screen "0017_Home Screen" 1280x800, template "Navigation"
   on GenerateScreen: SetTag("NavScreenChange", 7)
   on ClearScreen: SetTag("NavScreenChange", 0)
   GraphicView "Alarm Indicator Pump1" at 416,472 size 25x21; Picture "AlarmState2"
      Visibility <- "DB613_Komponent_State_GroupStatus{1}_FaultExist"
   GraphicView "Alarm Indicator Pump2" at 584,472 size 25x21; Picture "AlarmState2"
      Visibility <- "DB613_Komponent_State_GroupStatus{2}_FaultExist"
   GraphicView "Alarm Indicator hydraulic" at 1105,597 size 25x21; Picture "AlarmState2"
      Visibility <- "DB611_Hydraulic_State_MH_Hydraulic{1}_Fault_Exist"
   GraphicView "Alarm Indicator Pump2_1" at 508,688 size 25x21; Picture "AlarmState2"
      Visibility <- "DB614_MH_State_FaulExist"
   Button "Button_25" at 377,130 size 153x214; TextOff 'Text'; PictureOff "motor2"
      on Press: ActivateScreen("0006_Tank", 0); SetTag("DB612_Tank_State.ReadDeviceNo", 1); SetTag("NavScreenChange", 0)
   Button "Button_26" at 537,130 size 153x214; TextOff 'Text'; PictureOff "motor2"
      on Press: ActivateScreen("0006_Tank", 0); SetTag("DB612_Tank_State.ReadDeviceNo", 2); SetTag("NavScreenChange", 0)
   Button "b_Pump1" at 407,466 size 56x48; TextOff 'Text'
      on Press: ActivateScreen("0024_ActualFaults", 0); SetTag("Alarm_Filter_Tag", 3)
      ObjectEnable <- "DB613_Komponent_State_GroupStatus{1}_FaultExist"
   Button "b_Pump2" at 574,466 size 56x48; TextOff 'Text'
      ObjectEnable <- "DB613_Komponent_State_GroupStatus{2}_FaultExist"
      on Press: ActivateScreen("0024_ActualFaults", 0); SetTag("Alarm_Filter_Tag", 3); SetTag("NavScreenChange", 0)
   Button "b_hydraulic" at 1096,592 size 56x48; TextOff 'Text'
      on Press: ActivateScreen("0024_ActualFaults", 0); SetTag("Alarm_Filter_Tag", 2); SetTag("NavScreenChange", 0)
      ObjectEnable <- "DB611_Hydraulic_State_MH_Hydraulic{1}_Fault_Exist"
   Button "b_Pump2_1" at 494,677 size 56x48; TextOff 'Text'
      on Press: ActivateScreen("0024_ActualFaults", 0); SetTag("Alarm_Filter_Tag", 1); SetTag("NavScreenChange", 0)
      ObjectEnable <- "DB614_MH_State_FaulExist"
      Visibility <- "DB614_MH_State_FaulExist"
   GraphicView "Alarm Indicator Tank1" at 444,213 size 25x21; Picture "AlarmState2"
      Visibility <- "DB612_Tank_State_FaultExists{1}"
   GraphicView "Alarm Indicator Tank2" at 602,209 size 25x21; Picture "AlarmState2"
      Visibility <- "DB612_Tank_State_FaultExists{2}"
   Button "b_Tank1" at 432,208 size 50x36; TextOff 'Text'
      ObjectEnable <- "DB612_Tank_State_FaultExists{1}"
      on Press: ActivateScreen("0024_ActualFaults", 0); SetTag("Alarm_Filter_Tag", 4); SetTag("NavScreenChange", 0)
   Button "b_Tank2" at 588,208 size 50x36; TextOff 'Text'
      on Press: ActivateScreen("0024_ActualFaults", 0); SetTag("Alarm_Filter_Tag", 4); SetTag("NavScreenChange", 0)
      ObjectEnable <- "DB612_Tank_State_FaultExists{2}"
   TextField "Text field_8" at 549,392 size 129x30; Text '%'
      Visibility <- "DB702_Tank_Value_Tank{2}_With_Level_Probe"
   TextField "Text field_3" at 549,357 size 129x30; Text 'ºC'
   TextField "Text field_10" at 548,590 size 129x30; Text '%'
   TextField "Text field_14" at 548,526 size 129x30; Text 'bar'
   TextField "Text field_12" at 548,558 size 129x30; Text 'g/s'
   TextField "Text field_15" at 389,526 size 129x30; Text 'bar'
   TextField "Text field_9" at 389,590 size 129x30; Text '%'
   TextField "Text field_13" at 389,558 size 129x30; Text 'g/s'
   TextField "Text field_16" at 501,754 size 95x33; Text 'NL'
      Visibility <- "DB704_MH_Value_Mixinghead{0}_WithInerting"
   TextField "Text field_7" at 389,392 size 129x30; Text '%'
      Visibility <- "DB702_Tank_Value_Tank{1}_With_Level_Probe"
   TextField "Text field_4" at 389,357 size 129x30; Text 'ºC'
   TextField "Text field_2" at 595,640 size 95x33; Text 'bar'
   TextField "Text field_1" at 594,677 size 95x33; Text 'ºC'
   TextField "Text field_6" at 375,677 size 95x33; Text 'ºC'
   IOField "I/O field_20" at 501,754 size 73x33; FormatPattern 9999.9
      ProcessValue <- "DB619_State_MPart_ActMHInerting{1}_Total_Flow_N2_Visu"
      Visibility <- "DB704_MH_Value_Mixinghead{0}_WithInerting"
   IOField "I/O field_11" at 389,357 size 93x30; FormatPattern 9999.9
      ProcessValue <- "DB602_PV_Tank_Tank{1}_Temp_PV_ActV_Value"
   IOField "I/O field_12" at 549,357 size 93x30; FormatPattern 9999.9
      ProcessValue <- "DB602_PV_Tank_Tank{2}_Temp_PV_ActV_Value"
   IOField "I/O field_3" at 595,640 size 73x33; FormatPattern 9999.9
      ProcessValue <- "DB619_State_MPart_ActMHPressureMa{1}_Comp{2}"
   GraphicView "Graphic view_1" at 387,128 size 129x217; Picture "tank"
   GraphicView "Graphic view_2" at 549,128 size 129x217; Picture "tank"
   Button "Button_19" at 391,468 size 121x46; TextOff 'Text'; PictureOff "motor"
      on Click: SetTag("DB613_Komponent_State_ReadDeviceNo", 1); SetTag("NavScreenChange", 0); ActivateScreen("0010_Pump", 0)
   Button "Button_20" at 552,468 size 121x46; TextOff 'Text'; PictureOff "motor2"
      on Click: SetTag("DB613_Komponent_State_ReadDeviceNo", 2); SetTag("NavScreenChange", 0); ActivateScreen("0010_Pump", 0)
   Button "Button_22" at 987,418 size 162x134; TextOff 'MACHINE'; PictureOff "Machine"
      on Press: ActivateScreen("0021_Machine", 0); SetTag("NavScreenChange", 0)
   IOField "I/O field_43" at 378,97 size 151x30; FormatPattern ????????????????????
      ProcessValue <- "DB702_Tank_Value_Tank{1}_Name"
      Appearance <- "DB702_Tank_Value_Tank{1}_Color"
   IOField "I/O field_13" at 538,97 size 151x30; FormatPattern ????????????????????
      Appearance <- "DB702_Tank_Value_Tank{2}_Color"
      ProcessValue <- "DB702_Tank_Value_Tank{2}_Name"
   IOField "I/O field_14" at 378,426 size 151x30; FormatPattern ????????????????????
      Appearance <- "DB702_Tank_Value_Tank{1}_Color"
      ProcessValue <- "DB753_MeteringPump_Pump{1}_Name"
   IOField "I/O field_15" at 538,426 size 151x30; FormatPattern ????????????????????
      Appearance <- "DB702_Tank_Value_Tank{2}_Color"
      ProcessValue <- "DB753_MeteringPump_Pump{2}_Name"
   IOField "I/O field_16" at 703,651 size 151x30; FormatPattern ????????????????????
      Appearance <- "DB702_Tank_Value_Tank{2}_Color"
      ProcessValue <- "DB753_MeteringPump_Pump{2}_Name"
   IOField "I/O field_17" at 212,651 size 151x30; FormatPattern ????????????????????
      ProcessValue <- "DB753_MeteringPump_Pump{1}_Name"
      Appearance <- "DB702_Tank_Value_Tank{1}_Color"
   Button "Button_3" at 1015,579 size 139x135; TextOff 'MH hydrlc'; PictureOff "Mcn"
      on Press: ActivateScreen("0002_MixingHeadHydraulic", 0); SetTag("NavScreenChange", 0)
   TextField "Text field_11" at 459,754 size 41x33; Text 'N2'
      Visibility <- "DB704_MH_Value_Mixinghead{0}_WithInerting"
   GraphicView "Graphic view_3" at 478,640 size 104x112; Picture "images_4"
   GraphicView "Graphic view_5" at 483,637 size 28x27; Picture "cp2"
      Visibility <- "DB614_MH_State_MH_CleaningPiston{0}_Switch_CP_Forward"
   Bar "Bar_2" at 598,166 size 33x142; MinimumValue 0; MaximumValue 100
      ProcessValue <- "DB602_PV_Tank_Tank{2}_Level_PV_ActV_Value"
   TextField "Text field_5" at 375,640 size 95x33; Text 'bar'
   IOField "I/O field_4" at 376,677 size 73x33; FormatPattern 9999.9
      ProcessValue <- "DB619_State_MPart_ActMHTemperatureMa{1}_Comp{1}"
   IOField "I/O field_18" at 389,392 size 93x30; FormatPattern 9999.9
      ProcessValue <- "DB602_PV_Tank_Tank{1}_Level_PV_ActV_Value"
      Visibility <- "DB702_Tank_Value_Tank{1}_With_Level_Probe"
   IOField "I/O field_1" at 594,677 size 73x33; FormatPattern 9999.9
      ProcessValue <- "DB619_State_MPart_ActMHTemperatureMa{1}_Comp{2}"
   IOField "I/O field_19" at 549,392 size 93x30; FormatPattern 9999.9
      ProcessValue <- "DB602_PV_Tank_Tank{2}_Level_PV_ActV_Value"
      Visibility <- "DB702_Tank_Value_Tank{2}_With_Level_Probe"
   IOField "I/O field_5" at 389,526 size 97x30; FormatPattern 9999.9
      ProcessValue <- "DB608_PV_Metering_Metering{1}_Pressure_PV_ActV_Value"
   IOField "I/O field_7" at 548,526 size 97x30; FormatPattern 9999.9
      ProcessValue <- "DB608_PV_Metering_Metering{2}_Pressure_PV_ActV_Value"
   IOField "I/O field_8" at 548,558 size 97x30; FormatPattern 9999.99
      ProcessValue <- "DB608_PV_Metering_Metering{2}_Flow_PV_ActV_Value"
   IOField "I/O field_6" at 389,558 size 97x30; FormatPattern 9999.99
      ProcessValue <- "DB608_PV_Metering_Metering{1}_Flow_PV_ActV_Value"
   IOField "I/O field_9" at 389,590 size 97x30; FormatPattern 9999.9
      ProcessValue <- "DB608_PV_Metering_Metering{1}_MixingRatio_PV_ActV_Value"
   SymbolicIOField "Symbolic I/O field_1" at 406,718 size 102x33; TextOff '0'; TextOn '1'; TextList "MH_NO"
      ProcessValue <- "DB619_State_MPart_SWU{1}_ActualSWU"
      Visibility <- "DB619_State_MPart_SWU{1}_ActualSWU"
   Button "Button_21" at 479,637 size 104x112; TextOff 'Mixinghead'
      on Click: ActivateScreen("0004_Mixinghead", 0)
   IOField "I/O field_10" at 548,590 size 97x30; FormatPattern 9999.9
      ProcessValue <- "DB608_PV_Metering_Metering{2}_MixingRatio_PV_ActV_Value"
   Button "Button_2" at 543,522 size 140x103; TextOff 'Text'
      on Click: SetTag("DB613_Komponent_State_ReadDeviceNo", 2); SetTag("NavScreenChange", 0); ActivateScreen("0010_Pump", 0)
   Button "Button_1" at 383,522 size 140x102; TextOff 'Text'
      on Click: SetTag("DB613_Komponent_State_ReadDeviceNo", 1); SetTag("NavScreenChange", 0); ActivateScreen("0010_Pump", 0)
   GraphicView "ABB ROBOT" at 965,109 size 198x244; Picture "ABB Robot"
      Visibility <- "DB1901_Config_Robots_Config_Robots{0}_Type_ABB"
   GraphicView "KUKA ROBOT" at 965,109 size 198x244; Picture "Kuka Robot"
      Visibility <- "DB1901_Config_Robots_Config_Robots{0}_Type_Kuka"
   GraphicView "MOTOMAN ROBOT" at 965,109 size 198x244; Picture "Motoman Robot"
      Visibility <- "DB1901_Config_Robots_Config_Robots{0}_Type_Motoman"
   GraphicView "FANUC ROBOT" at 965,109 size 198x244; Picture "Fanuc Robot"
      Visibility <- "DB1901_Config_Robots_Config_Robots{0}_Type_Fanuc"
   Button "Button_27" at 955,97 size 175x267; TextOff 'Robot'
      on Click: ActivateScreen("0034_Robot", 0)
      Visibility <- "DB704_MH_Value_Mixinghead{0}_Conf_IntWithRobot"
   IOField "I/O field_2" at 375,640 size 73x33; FormatPattern 9999.9
      ProcessValue <- "DB619_State_MPart_ActMHPressureMa{1}_Comp{1}"
   Rectangle "Rectangle_8" at 598,166 size 33x142
      Visibility <- "DB612_Tank_State_Tank{2}_Max_Level"
   Rectangle "Rectangle_3" at 598,262 size 33x46
      Visibility <- "DB612_Tank_State_Tank{2}_Min_Level"
   Rectangle "Rectangle_5" at 598,166 size 33x142
      Visibility <- "DB612_Tank_State_Tank{2}_Start_Level_Filling"
   Rectangle "Rectangle_4" at 598,166 size 33x142
      Visibility <- "DB612_Tank_State_Tank{2}_Max_Level"
   Rectangle "Rectangle_7" at 440,166 size 33x142
      Visibility <- "DB612_Tank_State_Tank{1}_Max_Level"
   Rectangle "Rectangle_2" at 440,262 size 33x46
      Visibility <- "DB612_Tank_State_Tank{1}_Min_Level"
   Rectangle "Rectangle_6" at 440,166 size 33x142
      Visibility <- "DB612_Tank_State_Tank{1}_Start_Level_Filling"
   Rectangle "Rectangle_1" at 440,166 size 33x142
      Visibility <- "DB612_Tank_State_Tank{1}_Max_Level"

screen "0002_MixingHeadHydraulic" 1280x800, template "Navigation"
   on GenerateScreen: SetBit("DB611_Hydraulic_State_Read"); SetTag("Navigation_7", 5)
   IOField "I/O field_1" at 782,261 size 81x30; Authorization "Operate"; FormatPattern 99999
      ProcessValue <- "DB721_MH_Hydraulic_MH_Hyd{0}_Hyd_P_Startup"
   IOField "I/O field_2" at 782,293 size 81x30; Authorization "Operate"; FormatPattern 99999
      ProcessValue <- "DB721_MH_Hydraulic_MH_Hyd{0}_Hyd_P_Supervision"
   IOField "I/O field_3" at 782,353 size 81x30; Authorization "Operate"; FormatPattern 99999
      ProcessValue <- "DB721_MH_Hydraulic_MH_Hyd{0}_Hyd_CP_Time"
   IOField "I/O field_4" at 782,385 size 81x30; Authorization "Operate"; FormatPattern 99999
      ProcessValue <- "DB721_MH_Hydraulic_MH_Hyd{0}_Hyd_SwitchOFFDelay"
   IOField "I/O field_5" at 782,417 size 81x30; Authorization "Operate"; FormatPattern 99999
      ProcessValue <- "DB721_MH_Hydraulic_MH_Hyd{0}_Hyd_PressureSwitch"
   IOField "I/O field_6" at 229,521 size 131x30; FormatPattern 9999
      ProcessValue <- "DB611_Hydraulic_State_MH_Hydraulic{0}_HourCounter"
   TextField "Text field_1" at 504,263 size 186x25; Text 'Built up time start:'
   TextField "Text field_2" at 504,295 size 233x25; Text 'Built up time operaring:'
   TextField "Text field_3" at 504,355 size 225x25; Text 'Pressuring time for CP:'
   TextField "Text field_4" at 504,387 size 144x25; Text 'Stand by time:'
   TextField "Text field_5" at 504,419 size 161x25; Text 'Pressuring time:'
   TextField "Text field_6" at 874,263 size 46x25; Text 's'
   TextField "Text field_7" at 874,295 size 46x25; Text 's'
   TextField "Text field_8" at 874,355 size 46x25; Text 's'
   TextField "Text field_9" at 874,387 size 46x25; Text 's'
   TextField "Text field_10" at 874,419 size 46x25; Text 's'
   TextField "Text field_11" at 362,523 size 46x25; Text 'h'
   TextField "Text field_12" at 493,497 size 79x25; Text 'Options'
      Visibility <- "MixingHead Options"
   TextField "Text field_13" at 493,530 size 220x25; Text 'With 2 press switches:'
      Visibility <- "MixingHead Options"
   TextField "Text field_14" at 493,557 size 64x25; Text 'spare:'
      Visibility <- "MixingHead Options"
   TextField "Text field_15" at 493,587 size 64x25; Text 'spare:'
      Visibility <- "MixingHead Options"
   TextField "Text field_16" at 493,617 size 64x25; Text 'spare:'
      Visibility <- "MixingHead Options"
   TextField "Text field_17" at 493,647 size 64x25; Text 'spare:'
      Visibility <- "MixingHead Options"
   GraphicView "Graphic view_4" at 111,179 size 250x272; Picture "Mcn"
   Button "Button_3" at 326,104 size 451x32; TextOff 'MixingHead Hydraulic'
   Button "Button_1" at 482,240 size 423x221; TextOff 'Text'
   Button "Button_2" at 481,468 size 423x220; TextOff 'Text'
      Visibility <- "MixingHead Options"
   Button "check_with_2_press_switch" at 829,527 size 45x30; TextOff 'Text'; PictureOff "download"; PictureList "Check_Uncheck"
      ProcessValue <- "DB721_MH_Hydraulic_Option{0}_With2PSwitch"
      Visibility <- "MixingHead Options"
      on Click: InvertBit("DB721_MH_Hydraulic_Option{0}_With2PSwitch")
   Button "b_Close_MHhydraulic" at 848,470 size 51x41; TextOff 'Text'; PictureOff "images (1)"
      Visibility <- "MixingHead Options"
      on Click: SetTag("MixingHead Options", 0); SetTag("NavScreenChange", 0)
   Button "Button_10" at 1006,248 size 81x116; TextOff 'Text'
   GraphicView "Graphic view_1" at 1019,305 size 55x55; Picture "H"
   Rectangle "Rectangle_1" at 1015,256 size 64x56
      Appearance <- "DB611_Hydraulic_State_MH_Hydraulic{0}_State_Hydraulic"
   GraphicIOField "Graphic I/O field_1" at 1023,260 size 48x48; PictureList "ON_OFF_SWITCH"
      ProcessValue <- "DB611_Hydraulic_State_MH_Hydraulic{0}_Switch_Hydraulic_ON_OFF"
   Button "Button_18" at 1002,240 size 88x128; TextOff 'Text'
      on Click: InvertBit("DB611_Hydraulic_State_MH_Hydraulic{0}_Switch_Hydraulic_ON_OFF")
   GraphicView "Graphic view_2" at 143,508 size 77x51; Picture "counter hydraulic"
   Button "Button_4" at 217,210 size 80x52; TextOff 'Text'
   GraphicView "Graphic view_3" at 250,224 size 25x25; Picture "AlarmState2"
      Visibility <- "DB611_Hydraulic_State_MH_Hydraulic{0}_Fault_Exist"
   Button "b_MH_Increase" at 789,104 size 46x32; TextOff 'Text'; PictureOff "right arrow"
   Button "b_MH_Decrease" at 267,104 size 46x32; TextOff 'Text'; PictureOff "left arrow"
   Button "Template_Button_41" at 16,724 size 68x66; TextOff 'Text'; PictureList "Ico_navigation_2"; PictureOff "Setting_Nav_7"; Authorization "User administration"
      ProcessValue <- "Nav_7"
      Visibility <- "NavUserChange"
      on Click: SetTag("MixingHead Options", 1)

screen "0024_ActualFaults" 1280x800, template "Navigation"
   on ClearScreen: SetTag("refresh_Alarm", 0); SetTag("NavScreenChange", 0)
   on GenerateScreen: SetTag("NavScreenChange", 1)
   AlarmView "Machine Display alarm" at 103,169 size 1072x522
      Visibility <- "Alarm_Filter_Tag"
   Button "Button_3" at 326,104 size 451x32; TextOff 'Actual Fault'; TextList "Alarm_Screen_Filter"
      ProcessValue <- "Alarm_Filter_Tag"
   Button "b_Actual_Alarm" at 1097,92 size 60x60; TextOff 'ACTUAL'; PictureOff "Graphic_28"
      Appearance <- "Alarm_Filter_Tag"
      on Press: SetTag("Alarm_Filter_Tag", 0)
   Button "b_ArchiveAlarm" at 1028,91 size 60x60; TextOff 'ARCHIV'; PictureOff "archiveFoam_1"
      on Click: SetTag("Alarm_Filter_Tag", 10)
      Visibility <- "Alarm_Filter_Tag"
   Button "b_System" at 799,712 size 60x60; TextOff 'System'; PictureOff "system messages"; PictureList "ico_System_message_2"
      Visibility <- "Alarm_Filter_Tag"
      Appearance <- "Alarm_Filter_Tag"
      on Click: SetTag("Alarm_Filter_Tag", 13)
      ProcessValue <- "Alarm_Filter_Tag"
   Button "b_Foaming" at 891,712 size 60x60; TextOff 'Foaming'; PictureList "ico_Foaming_2"
      Visibility <- "Alarm_Filter_Tag"
      Appearance <- "Alarm_Filter_Tag"
      on Click: SetTag("Alarm_Filter_Tag", 12)
      ProcessValue <- "Alarm_Filter_Tag"
   Button "b_FaultFoam" at 984,712 size 60x60; TextOff 'Fault/ Foam'; PictureList "ico_ActualFault_Foaming_2"
      on Click: SetTag("Alarm_Filter_Tag", 10)
      Visibility <- "Alarm_Filter_Tag"
      Appearance <- "Alarm_Filter_Tag"
      ProcessValue <- "Alarm_Filter_Tag"
   Button "b_USB" at 705,712 size 60x60; TextOff 'Export USB'; PictureOff "USB_1"
      on Click: function_e9be9208(1, "Schicht0", '\Storage Card USB\', 0)
   Button "b_Fault_1" at 1077,712 size 60x60; TextOff 'Fault'; PictureList "ico_Actual_Fault_2"
      on Click: SetTag("Alarm_Filter_Tag", 11)
      Visibility <- "Alarm_Filter_Tag"
      ProcessValue <- "Alarm_Filter_Tag"
      Appearance <- "Alarm_Filter_Tag"
   Button "b_Fault_2" at 1077,712 size 60x60; TextOff 'Fault'
      on Click: SetTag("Alarm_Filter_Tag", 11)
      Visibility <- "Alarm_Filter_Tag"
      Appearance <- "Alarm_Filter_Tag"
   Button "b_Foaming_1" at 891,712 size 60x60; TextOff 'Foaming'
      on Click: SetTag("Alarm_Filter_Tag", 12)
      Appearance <- "Alarm_Filter_Tag"
      Visibility <- "Alarm_Filter_Tag"
   Button "b_FaultFoam_1" at 984,712 size 60x60; TextOff 'Fault/ Foam'
      on Click: SetTag("Alarm_Filter_Tag", 10)
      Visibility <- "Alarm_Filter_Tag"
      Appearance <- "Alarm_Filter_Tag"
   Button "b_System_1" at 799,712 size 60x60; TextOff 'System'; PictureOff "system messages"
      on Click: SetTag("Alarm_Filter_Tag", 13)
      Appearance <- "Alarm_Filter_Tag"
      Visibility <- "Alarm_Filter_Tag"
   Button "b_ArchiveAlarm_1" at 1028,91 size 60x60; TextOff 'ARCHIV'; PictureOff "archiveFoam_2"
      on Click: SetTag("Alarm_Filter_Tag", 10)
      Visibility <- "Alarm_Filter_Tag"
   AlarmView "MixingHydraulic Display Alarm" at 103,169 size 1072x522
      Visibility <- "Alarm_Filter_Tag"
   AlarmView "Tank Display Alarm" at 103,169 size 1072x522
      Visibility <- "Alarm_Filter_Tag"
   AlarmView "Pump Display Alarm" at 103,169 size 1072x522
      Visibility <- "Alarm_Filter_Tag"
   AlarmView "Archive faults" at 103,169 size 1072x522; AlarmLog "Schicht0"
      Visibility <- "Alarm_Filter_Tag"
   AlarmView "Archive faults/foaming" at 103,169 size 1072x522; AlarmLog "Schicht0"
      Visibility <- "Alarm_Filter_Tag"
   AlarmView "Archive foaming data" at 103,169 size 1072x522; AlarmLog "Schicht0"
      Visibility <- "Alarm_Filter_Tag"
   AlarmView "Archive system message" at 103,169 size 1072x522; AlarmLog "Schicht0"
      Visibility <- "Alarm_Filter_Tag"
   Button "b_Alarm_MHhydraulic_1" at 122,712 size 60x60; TextOff 'Text'; PictureList "icon_MHalarm"
      Visibility <- "Alarm_Filter_Tag"
      ProcessValue <- "Alarm_Filter_Tag"
      Appearance <- "Alarm_Filter_Tag"
   AlarmView "MixingHead Display Alarm" at 103,169 size 1072x522
      Visibility <- "Alarm_Filter_Tag"
   Button "b_Alarm_MH" at 117,704 size 71x77; TextOff 'MH'
      on Press: SetTag("Alarm_Filter_Tag", 1)
      Visibility <- "Alarm_Filter_Tag"
   AlarmView "Current Display Alarm" at 103,169 size 1072x522
      Visibility <- "Alarm_Filter_Tag"
   Button "b_Alarm_MHhydraulic_2" at 210,712 size 60x60; TextOff 'Text'; PictureList "icon_MHhyraulic"
      Visibility <- "Alarm_Filter_Tag"
      Appearance <- "Alarm_Filter_Tag"
      ProcessValue <- "Alarm_Filter_Tag"
   Button "b_Alarm_MHhydraulic" at 205,704 size 71x77; TextOff 'HYDRLC'
      on Press: SetTag("Alarm_Filter_Tag", 2)
      Visibility <- "Alarm_Filter_Tag"
   Button "b_Alarm_MHhydraulic_3" at 297,712 size 60x60; TextOff 'Text'; PictureList "ico_Pump"
      Visibility <- "Alarm_Filter_Tag"
      Appearance <- "Alarm_Filter_Tag"
      ProcessValue <- "Alarm_Filter_Tag"
   Button "b_MH_DosingPump" at 292,704 size 71x77; TextOff 'DOSING'
      on Press: SetTag("Alarm_Filter_Tag", 3)
      Visibility <- "Alarm_Filter_Tag"
   Button "b_Alarm_MHhydraulic_4" at 471,712 size 60x60; TextOff 'Text'; PictureList "ico_machine"
      Visibility <- "Alarm_Filter_Tag"
      Appearance <- "Alarm_Filter_Tag"
      ProcessValue <- "Alarm_Filter_Tag"
   Button "b_Alarm_Machine" at 466,704 size 71x77; TextOff 'MCHN'
      on Press: SetTag("Alarm_Filter_Tag", 5)
      Visibility <- "Alarm_Filter_Tag"
   Button "b_Alarm_MHhydraulic_5" at 384,712 size 60x60; TextOff 'Text'; PictureList "ico_tank"
      Visibility <- "Alarm_Filter_Tag"
      Appearance <- "Alarm_Filter_Tag"
      ProcessValue <- "Alarm_Filter_Tag"
   Button "b_Alarm_Tank" at 379,704 size 71x77; TextOff 'TANK'
      on Press: SetTag("Alarm_Filter_Tag", 4)
      Visibility <- "Alarm_Filter_Tag"

screen "0015_Oscilloscope" 1280x800, template "Navigation"
   Button "Button_3" at 326,104 size 451x32; TextOff 'Oscilloscope'
   TrendView "Trend view_1" at 105,152 size 1067x565
      ValueAxis1Begin <- "DB025_Oszilloskop_SkalierungGraphLinks_Startwert"
      ValueAxis1End <- "DB025_Oszilloskop_SkalierungGraphLinks_Ebdwert"
      ValueAxis2Begin <- "DB025_Oszilloskop_SkalierungGraphRechts_Startwert"
      ValueAxis2End <- "DB025_Oszilloskop_SkalierungGraphRechts_Ebdwert"
   Button "Button_2" at 115,748 size 52x37; TextOff 'Text'; PictureOff "Graphic_32"
      on Click: function_e0f5d53a("Trend view_1")
   Button "Button_4" at 183,748 size 52x37; TextOff 'Text'; PictureOff "Graphic_31"
      on Click: function_e0f5d53a("Trend view_1")
   Button "Button_5" at 252,748 size 52x37; TextOff 'Text'; PictureOff "Graphic_33"
      on Click: function_b4e726f8("Trend view_1")
   Button "Button_6" at 320,748 size 52x37; TextOff 'Text'; PictureOff "Graphic_34"
      on Click: function_f26ff0ec("Trend view_1")
   Button "Button_7" at 389,748 size 52x37; TextOff 'Text'; PictureOff "Graphic_35"
      on Click: function_c2ce674d("Trend view_1")
   Button "Button_8" at 457,748 size 52x37; TextOff 'Text'; PictureOff "Graphic_36"
      on Click: function_f48c2799("Trend view_1")
   Button "Button_9" at 526,748 size 52x37; TextOff 'Text'; PictureOff "Graphic_37"
      on Click: function_b22ecfcd("Trend view_1")
   Button "Button_10" at 595,748 size 52x37; TextOff 'Text'; PictureOff "gear_setting"
      on Click: ActivateScreen("0016_Osciloscope Setting", 0)
   Button "Button_11" at 979,748 size 52x37; TextOff 'Text'; PictureOff "Graphic_38"
      on Click: function_a3fbdc78("Trend view_1")
   Button "Button_1" at 1047,748 size 52x37; TextOff 'Text'; PictureOff "Graphic_39"
      on Click: function_a16a7cb4("Trend view_1")
   Button "Button_12" at 1115,748 size 52x37; TextOff 'Text'; PictureOff "Graphic_40"
      on Click: function_c7513061("Trend view_1")

screen "0100_LargeScalledValues" 1280x800, template "Navigation"
   Button "Button_2" at 115,466 size 1047x206; TextOff 'Text'
      Appearance <- "DB702_Tank_Value_Tank{2}_Color"
      Visibility <- "LargeScalleValues Control"
   IOField "I/O field_4" at 172,488 size 328x166; FormatPattern 999.9
      ProcessValue <- "DB608_PV_Metering_Metering{2}_Pressure_PV_ActV_Value"
      Visibility <- "LargeScalleValues Control"
   Button "Button_1" at 115,255 size 1047x206; TextOff 'Text'
      Appearance <- "DB702_Tank_Value_Tank{1}_Color"
      Visibility <- "LargeScalleValues Control"
   IOField "I/O field_1" at 172,280 size 328x166; FormatPattern 999.9
      ProcessValue <- "DB608_PV_Metering_Metering{1}_Pressure_PV_ActV_Value"
      Visibility <- "LargeScalleValues Control"
   IOField "I/O field_2" at 836,280 size 328x166; FormatPattern 999.9
      ProcessValue <- "DB608_PV_Metering_Metering{1}_Flow_PV_ActV_Value"
      Visibility <- "LargeScalleValues Control"
   IOField "I/O field_3" at 836,488 size 328x166; FormatPattern 999.9
      ProcessValue <- "DB608_PV_Metering_Metering{2}_Flow_PV_ActV_Value"
      Visibility <- "LargeScalleValues Control"
   TextField "Text field_1" at 252,132 size 192x120; Text 'bar'
      Visibility <- "LargeScalleValues Control"
   TextField "Text field_2" at 872,132 size 192x120; Text 'g/s'
      Visibility <- "LargeScalleValues Control"
   Button "Button_4" at 115,466 size 1047x206; TextOff 'Text'
      Appearance <- "DB702_Tank_Value_Tank{2}_Color"
      Visibility <- "LargeScalleValues Control"
   Button "Button_5" at 115,255 size 1047x206; TextOff 'Text'
      Appearance <- "DB702_Tank_Value_Tank{1}_Color"
      Visibility <- "LargeScalleValues Control"
   IOField "I/O field_5" at 479,280 size 328x166; FormatPattern 999.9
      ProcessValue <- "DB602_PV_Tank_Tank{1}_Level_PV_ActV_Value"
      Visibility <- "LargeScalleValues Control"
   IOField "I/O field_6" at 476,494 size 328x166; FormatPattern 999.9
      ProcessValue <- "DB602_PV_Tank_Tank{2}_Level_PV_ActV_Value"
      Visibility <- "LargeScalleValues Control"
   TextField "Text field_3" at 894,308 size 192x120; Text '%'
      Visibility <- "LargeScalleValues Control"
   TextField "Text field_7" at 894,509 size 192x120; Text '%'
      Visibility <- "LargeScalleValues Control"
   Button "Button_6" at 115,466 size 1047x206; TextOff 'Text'
      Visibility <- "LargeScalleValues Control"
      Appearance <- "DB702_Tank_Value_Tank{2}_Color"
   Button "Button_7" at 115,255 size 1047x206; TextOff 'Text'
      Appearance <- "DB702_Tank_Value_Tank{1}_Color"
      Visibility <- "LargeScalleValues Control"
   TextField "Text field_4" at 252,132 size 192x120; Text 'bar'
      Visibility <- "LargeScalleValues Control"
   TextField "Text field_5" at 872,132 size 192x120; Text 'g/s'
      Visibility <- "LargeScalleValues Control"
   IOField "I/O field_7" at 172,280 size 328x166; FormatPattern 999.9
      ProcessValue <- "DB619_State_MPart_ActMHPressureMa{1}_Comp{1}"
      Visibility <- "LargeScalleValues Control"
   IOField "I/O field_8" at 836,280 size 328x166; FormatPattern 999.9
      ProcessValue <- "DB608_PV_Metering_Metering{1}_Flow_PV_ActV_Value"
      Visibility <- "LargeScalleValues Control"
   IOField "I/O field_9" at 836,488 size 328x166; FormatPattern 999.9
      ProcessValue <- "DB608_PV_Metering_Metering{2}_Flow_PV_ActV_Value"
      Appearance <- "DB702_Tank_Value_Tank{2}_Color"
      Visibility <- "LargeScalleValues Control"
   IOField "I/O field_10" at 172,488 size 328x166; FormatPattern 999.9
      ProcessValue <- "DB619_State_MPart_ActMHPressureMa{1}_Comp{2}"
      Visibility <- "LargeScalleValues Control"
   TextField "Text field_6" at 447,132 size 383x120; Text '---'
      Visibility <- "LargeScalleValues Control"
   Button "Button_8" at 135,711 size 60x60; TextOff 'Text'; PictureList "ico_MH"
      Appearance <- "LargeScalleValues Control"
      ProcessValue <- "LargeScalleValues Control"
   Button "Button_3" at 326,104 size 451x32; TextOff 'Large Scalled Values'
   Button "Button_9" at 296,711 size 60x60; TextOff 'Text'; PictureOff "tank"
      Appearance <- "LargeScalleValues Control"
   Button "Button_10" at 216,711 size 60x60; TextOff 'Text'; PictureOff "Graphic_1"; PictureList "ico_Pump_large"
      Appearance <- "LargeScalleValues Control"
      ProcessValue <- "LargeScalleValues Control"
   Button "b_MH_large" at 135,711 size 60x60; TextOff 'MH'; PictureList "MixingHead"
      Appearance <- "LargeScalleValues Control"
      on Click: SetTag("LargeScalleValues Control", 0)
   Button "b_pump_" at 216,711 size 60x60; TextOff 'Tank'; PictureList "tank"
      on Click: SetTag("LargeScalleValues Control", 1)
   Button "b_tank_large_1" at 296,711 size 60x60; TextOff 'Tank'; PictureList "tank"
      on Click: SetTag("LargeScalleValues Control", 2)
      Appearance <- "LargeScalleValues Control"

screen "0009_Switch Menu" 1280x800, template "Navigation"
   Button "Button_1" at 164,321 size 430x30; TextOff 'Text'
      Appearance <- "DB702_Tank_Value_Tank{1}_Color"
   Button "Button_2" at 646,322 size 432x30; TextOff 'Text'
      Appearance <- "DB702_Tank_Value_Tank{2}_Color"
   Button "Button_3" at 326,104 size 451x32; TextOff 'Switch Menu'
   Button "Button_5" at 164,376 size 81x116; TextOff 'Text'
      Visibility <- "DB702_Tank_Value_Tank{1}_With_Tempering_Heizung"
   Button "Button_4" at 252,376 size 81x116; TextOff 'Text'
      Visibility <- "DB702_Tank_Value_Tank{1}_With_Filling"
   Button "Button_6" at 340,376 size 81x116; TextOff 'Text'
      Visibility <- "DB702_Tank_Value_Tank{1}_With_Agitator"
   Button "Button_7" at 648,376 size 81x116; TextOff 'Text'
      Visibility <- "DB702_Tank_Value_Tank{2}_With_Tempering_Heizung"
   Button "Button_8" at 736,376 size 81x116; TextOff 'Text'
      Visibility <- "DB702_Tank_Value_Tank{2}_With_Filling"
   Button "Button_9" at 824,376 size 81x116; TextOff 'Text'
      Visibility <- "DB702_Tank_Value_Tank{2}_With_Agitator"
   Button "Button_10" at 165,160 size 81x116; TextOff 'Text'
   Button "Button_11" at 253,160 size 81x116; TextOff 'Text'
   Button "Button_12" at 341,160 size 81x116; TextOff 'Text'
   Button "Button_13" at 429,160 size 81x116; TextOff 'Text'
   Button "Button_14" at 428,375 size 81x116; TextOff 'Text'
      Visibility <- "DB753_MeteringPump_Pump{1}_WithEdgeFilter"
   Button "Button_15" at 516,374 size 81x116; TextOff 'Text'
      Visibility <- "DB753_MeteringPump_Pump{1}_WithHeating"
   Button "Button_16" at 911,376 size 81x116; TextOff 'Text'
      Visibility <- "DB753_MeteringPump_Pump{2}_WithEdgeFilter"
   Button "Button_17" at 997,376 size 81x116; TextOff 'Text'
      Visibility <- "DB753_MeteringPump_Pump{2}_WithHeating"
   GraphicView "Graphic view_1" at 178,218 size 55x55; Picture "H"
   GraphicView "Graphic view_2" at 270,222 size 48x48; Picture "REDUCED"
   GraphicView "Graphic view_3" at 359,222 size 48x48; Picture "Interval"
   GraphicView "Graphic view_4" at 446,222 size 48x48; Picture "LowPress"
   GraphicView "Graphic view_5" at 176,441 size 56x48; Picture "Switch Temp"
      Visibility <- "DB702_Tank_Value_Tank{1}_With_Tempering_Heizung"
   GraphicView "Graphic view_6" at 264,440 size 56x48; Picture "Refilling"
      Visibility <- "DB702_Tank_Value_Tank{1}_With_Filling"
   GraphicView "Graphic view_7" at 352,440 size 56x48; Picture "Agitator"
      Visibility <- "DB702_Tank_Value_Tank{1}_With_Agitator"
   GraphicView "Graphic view_8" at 663,440 size 56x48; Picture "Switch Temp"
      Visibility <- "DB702_Tank_Value_Tank{2}_With_Tempering_Heizung"
   GraphicView "Graphic view_9" at 751,439 size 56x48; Picture "Refilling"
      Visibility <- "DB702_Tank_Value_Tank{2}_With_Filling"
   GraphicView "Graphic view_10" at 838,440 size 56x48; Picture "Agitator"
      Visibility <- "DB702_Tank_Value_Tank{2}_With_Agitator"
   Rectangle "Rectangle_1" at 174,168 size 64x56
      Appearance <- "DB611_Hydraulic_State_MH_Hydraulic{1}_State_Hydraulic"
   GraphicIOField "Graphic I/O field_1" at 182,172 size 48x48; PictureList "ON_OFF_SWITCH"
      ProcessValue <- "DB611_Hydraulic_State_MH_Hydraulic{1}_Switch_Hydraulic_ON_OFF"
   Rectangle "Rectangle_3" at 261,168 size 64x56
      Appearance <- "DB619_State_MPart_Recirculation{1}_State_Reduced"
   Rectangle "Rectangle_4" at 349,168 size 64x56
      Appearance <- "DB619_State_MPart_Recirculation{1}_State_Intervall"
   GraphicIOField "Graphic I/O field_2" at 269,171 size 48x48; PictureList "ON_OFF_SWITCH"
      ProcessValue <- "DB619_State_MPart_Recirculation{1}_Switch_Reduced"
   GraphicIOField "Graphic I/O field_3" at 357,171 size 48x48; PictureList "ON_OFF_SWITCH"
      ProcessValue <- "DB619_State_MPart_Recirculation{1}_Switch_Intervall"
   Rectangle "Rectangle_5" at 437,168 size 64x56
      Appearance <- "DB619_State_MPart_Recirculation{1}_State_Lowpressure"
   GraphicIOField "Graphic I/O field_4" at 445,171 size 48x48; PictureList "ON_OFF_SWITCH"
      ProcessValue <- "DB619_State_MPart_Recirculation{1}_Switch_Lowpressure"
   Rectangle "Rectangle_6" at 173,384 size 64x56
      Appearance <- "DB612_Tank_State_ControllerTankTemp{1}_State_Temp"
      Visibility <- "DB702_Tank_Value_Tank{1}_With_Tempering_Heizung"
   Rectangle "Rectangle_7" at 260,384 size 64x56
      Appearance <- "DB612_Tank_State_Tank{1}_State_Refilling"
      Visibility <- "DB702_Tank_Value_Tank{1}_With_Filling"
   GraphicIOField "Graphic I/O field_5" at 181,387 size 48x48; PictureList "ON_OFF_SWITCH"
      ProcessValue <- "DB612_Tank_State_ControllerTankTemp{1}_Switch_Temp_ON_OFF"
      Visibility <- "DB702_Tank_Value_Tank{1}_With_Tempering_Heizung"
   GraphicIOField "Graphic I/O field_6" at 268,387 size 48x48; PictureList "ON_OFF_SWITCH"
      ProcessValue <- "DB612_Tank_State_Tank{1}_Switch_Refilling_ON_OFF"
      Visibility <- "DB702_Tank_Value_Tank{1}_With_Filling"
   Rectangle "Rectangle_8" at 349,384 size 64x56
      Appearance <- "DB612_Tank_State_Agitator{1}_State_Drive"
      Visibility <- "DB702_Tank_Value_Tank{1}_With_Agitator"
   GraphicIOField "Graphic I/O field_7" at 355,387 size 48x48; PictureList "ON_OFF_SWITCH"
      ProcessValue <- "DB612_Tank_State_Agitator{1}_Switch_Drive_ON_OFF"
      Visibility <- "DB702_Tank_Value_Tank{1}_With_Agitator"
   Rectangle "Rectangle_9" at 436,384 size 64x56
      Appearance <- "DB613_Komponent_State_EdgeFilter{1}_State_Drive"
      Visibility <- "DB753_MeteringPump_Pump{1}_WithEdgeFilter"
   GraphicIOField "Graphic I/O field_8" at 445,387 size 48x48; PictureList "ON_OFF_SWITCH"
      ProcessValue <- "DB613_Komponent_State_EdgeFilter{1}_Switch_Drive_ON_OFF"
      Visibility <- "DB753_MeteringPump_Pump{1}_WithEdgeFilter"
   Rectangle "Rectangle_10" at 525,384 size 64x56
      Appearance <- "DB613_Komponent_State_HeatexchangerHP{1}_State_Temp"
      Visibility <- "DB753_MeteringPump_Pump{1}_WithHeating"
   Rectangle "Rectangle_11" at 656,384 size 64x56
      Appearance <- "DB612_Tank_State_ControllerTankTemp{2}_State_Temp"
      Visibility <- "DB702_Tank_Value_Tank{2}_With_Tempering_Heizung"
   GraphicIOField "Graphic I/O field_9" at 533,387 size 48x48; PictureList "ON_OFF_SWITCH"
      ProcessValue <- "DB613_Komponent_State_HeatexchangerHP{1}_Switch_Temp_ON_OFF"
      Visibility <- "DB753_MeteringPump_Pump{1}_WithHeating"
   GraphicIOField "Graphic I/O field_10" at 664,387 size 48x48; PictureList "ON_OFF_SWITCH"
      ProcessValue <- "DB612_Tank_State_ControllerTankTemp{2}_Switch_Temp_ON_OFF"
      Visibility <- "DB702_Tank_Value_Tank{2}_With_Tempering_Heizung"
   Rectangle "Rectangle_12" at 745,384 size 64x56
      Appearance <- "DB612_Tank_State_Tank{2}_State_Refilling"
      Visibility <- "DB702_Tank_Value_Tank{2}_With_Filling"
   GraphicIOField "Graphic I/O field_11" at 753,387 size 48x48; PictureList "ON_OFF_SWITCH"
      ProcessValue <- "DB612_Tank_State_Tank{2}_Switch_Refilling_ON_OFF"
      Visibility <- "DB702_Tank_Value_Tank{2}_With_Filling"
   Rectangle "Rectangle_13" at 833,384 size 64x56
      Appearance <- "DB612_Tank_State_Agitator{2}_State_Drive"
      Visibility <- "DB702_Tank_Value_Tank{2}_With_Agitator"
   GraphicIOField "Graphic I/O field_12" at 841,387 size 48x48; PictureList "ON_OFF_SWITCH"
      ProcessValue <- "DB612_Tank_State_Agitator{2}_Switch_Drive_ON_OFF"
      Visibility <- "DB702_Tank_Value_Tank{2}_With_Agitator"
   Rectangle "Rectangle_14" at 920,384 size 64x56
      Appearance <- "DB613_Komponent_State_EdgeFilter{2}_State_Drive"
      Visibility <- "DB753_MeteringPump_Pump{2}_WithEdgeFilter"
   GraphicIOField "Graphic I/O field_13" at 928,387 size 48x48; PictureList "ON_OFF_SWITCH"
      ProcessValue <- "DB613_Komponent_State_EdgeFilter{2}_Switch_Drive_ON_OFF"
      Visibility <- "DB753_MeteringPump_Pump{2}_WithEdgeFilter"
   Rectangle "Rectangle_15" at 1006,384 size 64x56
      Appearance <- "DB613_Komponent_State_HeatexchangerHP{2}_State_Temp"
      Visibility <- "DB753_MeteringPump_Pump{2}_WithHeating"
   GraphicIOField "Graphic I/O field_14" at 1014,387 size 48x48; PictureList "ON_OFF_SWITCH"
      ProcessValue <- "DB613_Komponent_State_HeatexchangerHP{2}_Switch_Temp_ON_OFF"
      Visibility <- "DB753_MeteringPump_Pump{2}_WithHeating"
   Button "Button_32" at 163,506 size 81x116; TextOff 'Text'
      Visibility <- "DB753_MeteringPump_Pump{1}_WithLPHeatExchanger"
   Rectangle "Rectangle_16" at 172,516 size 64x56
      Appearance <- "DB613_Komponent_State_HeatexchangerLP{1}_State_Temp"
      Visibility <- "DB753_MeteringPump_Pump{1}_WithLPHeatExchanger"
   GraphicIOField "Graphic I/O field_15" at 180,519 size 48x48; PictureList "ON_OFF_SWITCH"
      ProcessValue <- "DB613_Komponent_State_HeatexchangerLP{1}_Switch_Temp_ON_OFF"
      Visibility <- "DB753_MeteringPump_Pump{1}_WithLPHeatExchanger"
   Button "Button_34" at 648,509 size 81x116; TextOff 'Text'
      Visibility <- "DB753_MeteringPump_Pump{2}_WithLPHeatExchanger"
   Rectangle "Rectangle_17" at 657,517 size 64x56
      Appearance <- "DB613_Komponent_State_HeatexchangerLP{2}_State_Temp"
      Visibility <- "DB753_MeteringPump_Pump{2}_WithLPHeatExchanger"
   GraphicIOField "Graphic I/O field_16" at 665,520 size 48x48; PictureList "ON_OFF_SWITCH"
      ProcessValue <- "DB613_Komponent_State_HeatexchangerLP{2}_Switch_Temp_ON_OFF"
      Visibility <- "DB753_MeteringPump_Pump{2}_WithLPHeatExchanger"
   GraphicView "Graphic view_11" at 444,442 size 44x43; Picture "edgefilter"
      Visibility <- "DB753_MeteringPump_Pump{1}_WithEdgeFilter"
   GraphicView "Graphic view_12" at 930,441 size 44x43; Picture "edgefilter"
      Visibility <- "DB753_MeteringPump_Pump{2}_WithEdgeFilter"
   GraphicView "Graphic view_13" at 518,442 size 79x52; Picture "SWITCH HEATHP"
      Visibility <- "DB753_MeteringPump_Pump{1}_WithHeating"
   GraphicView "Graphic view_14" at 997,442 size 79x52; Picture "SWITCH HEATHP"
      Visibility <- "DB753_MeteringPump_Pump{2}_WithHeating"
   GraphicView "Graphic view_15" at 165,573 size 76x43; Picture "Switch heatLP"
      Visibility <- "DB753_MeteringPump_Pump{1}_WithLPHeatExchanger"
   GraphicView "Graphic view_16" at 650,578 size 76x43; Picture "Switch heatLP"
      Visibility <- "DB753_MeteringPump_Pump{2}_WithLPHeatExchanger"
   Button "Button_36" at 647,160 size 81x116; TextOff 'Text'
      Visibility <- "DB790_PlantParameter_AmountMachine"
   Button "Button_37" at 735,160 size 81x116; TextOff 'Text'
      Visibility <- "DB790_PlantParameter_AmountMachine"
   Button "Button_38" at 823,160 size 81x116; TextOff 'Text'
      Visibility <- "DB790_PlantParameter_AmountMachine"
   Button "Button_39" at 911,160 size 81x116; TextOff 'Text'
      Visibility <- "DB790_PlantParameter_AmountMachine"
   GraphicView "Graphic view_17" at 660,218 size 55x55; Picture "H"
      Visibility <- "DB790_PlantParameter_AmountMachine"
   GraphicView "Graphic view_18" at 752,222 size 48x48; Picture "REDUCED"
      Visibility <- "DB790_PlantParameter_AmountMachine"
   GraphicView "Graphic view_19" at 841,222 size 48x48; Picture "Interval"
      Visibility <- "DB790_PlantParameter_AmountMachine"
   GraphicView "Graphic view_20" at 928,222 size 48x48; Picture "LowPress"
      Visibility <- "DB790_PlantParameter_AmountMachine"
   Rectangle "Rectangle_18" at 656,168 size 64x56
      Visibility <- "DB790_PlantParameter_AmountMachine"
      Appearance <- "DB611_Hydraulic_State_MH_Hydraulic{2}_State_Hydraulic"
   GraphicIOField "Graphic I/O field_17" at 664,172 size 48x48; PictureList "ON_OFF_SWITCH"
      Visibility <- "DB790_PlantParameter_AmountMachine"
      ProcessValue <- "DB611_Hydraulic_State_MH_Hydraulic{2}_Switch_Hydraulic_ON_OFF"
   Rectangle "Rectangle_19" at 743,168 size 64x56
      Visibility <- "DB790_PlantParameter_AmountMachine"
      Appearance <- "DB619_State_MPart_Recirculation{2}_State_Reduced"
   Rectangle "Rectangle_20" at 831,168 size 64x56
      Visibility <- "DB790_PlantParameter_AmountMachine"
      Appearance <- "DB619_State_MPart_Recirculation{2}_State_Intervall"
   GraphicIOField "Graphic I/O field_18" at 751,171 size 48x48; PictureList "ON_OFF_SWITCH"
      Visibility <- "DB790_PlantParameter_AmountMachine"
      ProcessValue <- "DB619_State_MPart_Recirculation{2}_Switch_Reduced"
   GraphicIOField "Graphic I/O field_19" at 839,171 size 48x48; PictureList "ON_OFF_SWITCH"
      Visibility <- "DB790_PlantParameter_AmountMachine"
      ProcessValue <- "DB619_State_MPart_Recirculation{2}_Switch_Intervall"
   Rectangle "Rectangle_21" at 919,168 size 64x56
      Visibility <- "DB790_PlantParameter_AmountMachine"
      Appearance <- "DB619_State_MPart_Recirculation{2}_State_Lowpressure"
   GraphicIOField "Graphic I/O field_20" at 927,171 size 48x48; PictureList "ON_OFF_SWITCH"
      Visibility <- "DB790_PlantParameter_AmountMachine"
      ProcessValue <- "DB619_State_MPart_Recirculation{2}_Switch_Lowpressure"
   Button "Button_18" at 161,152 size 88x128; TextOff 'Text'
      on Click: InvertBit("DB611_Hydraulic_State_MH_Hydraulic{1}_Switch_Hydraulic_ON_OFF")
   Button "Button_19" at 251,152 size 88x128; TextOff 'Text'
      on Click: InvertBit("DB619_State_MPart_Recirculation{1}_Switch_Reduced")
   Button "Button_20" at 336,152 size 88x128; TextOff 'Text'
      on Click: InvertBit("DB619_State_MPart_Recirculation{1}_Switch_Intervall")
   Button "Button_21" at 425,152 size 88x128; TextOff 'Text'
      on Click: InvertBit("DB619_State_MPart_Recirculation{1}_Switch_Lowpressure")
   Button "Button_40" at 643,152 size 88x128; TextOff 'Text'
      on Click: InvertBit("DB611_Hydraulic_State_MH_Hydraulic{2}_Switch_Hydraulic_ON_OFF")
      Visibility <- "DB790_PlantParameter_AmountMachine"
   Button "Button_41" at 733,152 size 88x128; TextOff 'Text'
      on Click: InvertBit("DB619_State_MPart_Recirculation{2}_Switch_Reduced")
      Visibility <- "DB790_PlantParameter_AmountMachine"
   Button "Button_42" at 818,152 size 88x128; TextOff 'Text'
      on Click: InvertBit("DB619_State_MPart_Recirculation{2}_Switch_Intervall")
      Visibility <- "DB790_PlantParameter_AmountMachine"
   Button "Button_43" at 907,152 size 88x128; TextOff 'Text'
      on Click: InvertBit("DB619_State_MPart_Recirculation{2}_Switch_Lowpressure")
      Visibility <- "DB790_PlantParameter_AmountMachine"
   Button "Button_31" at 992,368 size 88x128; TextOff 'Text'
      on Click: InvertBit("DB613_Komponent_State_HeatexchangerHP{2}_Switch_Temp_ON_OFF")
      Visibility <- "DB753_MeteringPump_Pump{2}_WithHeating"
   Button "Button_30" at 905,368 size 88x128; TextOff 'Text'
      on Click: InvertBit("DB613_Komponent_State_EdgeFilter{2}_Switch_Drive_ON_OFF")
      Visibility <- "DB753_MeteringPump_Pump{2}_WithEdgeFilter"
   Button "Button_29" at 818,368 size 88x128; TextOff 'Text'
      on Click: InvertBit("DB612_Tank_State_Agitator{2}_Switch_Drive_ON_OFF")
      Visibility <- "DB702_Tank_Value_Tank{2}_With_Agitator"
   Button "Button_28" at 731,368 size 88x128; TextOff 'Text'
      on Click: InvertBit("DB612_Tank_State_Tank{2}_Switch_Refilling_ON_OFF")
      Visibility <- "DB702_Tank_Value_Tank{2}_With_Filling"
   Button "Button_27" at 644,368 size 88x128; TextOff 'Text'
      on Click: InvertBit("DB612_Tank_State_ControllerTankTemp{2}_Switch_Temp_ON_OFF")
      Visibility <- "DB702_Tank_Value_Tank{2}_With_Tempering_Heizung"
   Button "Button_35" at 643,501 size 88x128; TextOff 'Text'
      on Click: InvertBit("DB613_Komponent_State_HeatexchangerLP{2}_Switch_Temp_ON_OFF")
      Visibility <- "DB753_MeteringPump_Pump{2}_WithLPHeatExchanger"
   Button "Button_26" at 513,368 size 88x128; TextOff 'Text'
      on Click: InvertBit("DB613_Komponent_State_HeatexchangerHP{1}_Switch_Temp_ON_OFF")
      Visibility <- "DB753_MeteringPump_Pump{1}_WithHeating"
   Button "Button_25" at 425,368 size 88x128; TextOff 'Text'
      on Click: InvertBit("DB613_Komponent_State_EdgeFilter{1}_Switch_Drive_ON_OFF")
      Visibility <- "DB753_MeteringPump_Pump{1}_WithEdgeFilter"
   Button "Button_24" at 338,368 size 88x128; TextOff 'Text'
      on Click: InvertBit("DB612_Tank_State_Agitator{1}_Switch_Drive_ON_OFF")
      Visibility <- "DB702_Tank_Value_Tank{1}_With_Agitator"
   Button "Button_23" at 249,368 size 88x128; TextOff 'Text'
      on Click: InvertBit("DB612_Tank_State_Tank{1}_Switch_Refilling_ON_OFF")
      Visibility <- "DB702_Tank_Value_Tank{1}_With_Filling"
   Button "Button_22" at 160,368 size 88x128; TextOff 'Text'
      on Click: InvertBit("DB612_Tank_State_ControllerTankTemp{1}_Switch_Temp_ON_OFF")
      Visibility <- "DB702_Tank_Value_Tank{1}_With_Tempering_Heizung"
   Button "Button_33" at 160,500 size 88x128; TextOff 'Text'
      on Click: InvertBit("DB613_Komponent_State_HeatexchangerLP{1}_Switch_Temp_ON_OFF")
      Visibility <- "DB753_MeteringPump_Pump{1}_WithLPHeatExchanger"

screen "0018_SystemSetting" 1280x800, template "Navigation"
   on GenerateScreen: SetTag("NavScreenChange", 2)
   on ClearScreen: SetTag("NavScreenChange", 0)
   Button "Button_3" at 326,104 size 451x32; TextOff 'System Settings'
   Button "b_print" at 592,704 size 60x60; TextOff 'Text'; PictureOff "printer off"
      Visibility <- "System Setting Screen Control"
      on Click: function_fd03fc5c("Shot Data"); InvertBit("Print Function")
   Button "b_setdatetime" at 881,704 size 60x60; TextOff 'Text'; PictureOff "datetime"
      on Press: function_efd93a16("Change DateTime", 300, 344, -1, -1, 1)
      Visibility <- "System Setting Screen Control"
   Button "b_calibration" at 978,703 size 60x60; TextOff 'Text'; PictureOff "touch"
      Visibility <- "System Setting Screen Control"
      on Click: function_bc3e350c()
   Button "b_cleanscreen" at 1072,703 size 60x60; TextOff 'Text'; PictureOff "paint"
      on Press: function_be740847(30)
      Visibility <- "System Setting Screen Control"
   Button "b_setting" at 248,704 size 60x60; TextOff 'Text'; PictureOff "Setting_Nav_7"; Authorization "User administration"
      Visibility <- "System Setting Screen Control"
      on Click: function_f34a74f3()
   Button "b_logout" at 784,704 size 60x60; TextOff 'Text'; PictureOff "logoff"
      on Press: function_f23ef4c9()
      Visibility <- "System Setting Screen Control"
   Button "b_networksetting" at 495,704 size 60x60; TextOff 'Text'; PictureOff "ethernet"
      on Click: ActivateScreen("0014_Network Setting", 0)
      Visibility <- "NavUserChange"
   Button "b_Stop" at 153,704 size 60x60; TextOff 'Stop Runtime'; PictureOff "door"
      on Press: StopRuntime(0)
      Visibility <- "NavUserChange"
   UserView "User view_1" at 128,153 size 1032x520
   StatusForce "Watch table_1" at 137,173 size 1003x605; ToolTipText 'Text'
      Visibility <- "System Setting Screen Control"